(* Logix 5000 project; controller PLC_MCC1300_75F1 vendor 1 type 14 code 166 rev 32.11; software revision 32.04; part 64 of 83 *)
(* tags used below, declared in another part *)
   AUX_tConvoy_SL_NULL : UDT_Convoy_SL;
   CONST_rgdDestMask : DINT[32];   // Destination Mask
   CONST_tPlant : UDT_PLANT_CONSTANTS;
   GP_TrackingSearchPlate : GP_TrackingSearchPlate;
   M315Popup : MAC_Popup_ZC[2];
   M315Popup_HMW : MAC_Popup_ZC_HMW[2];
   M315Popup_ReentryCap : UDT_ConvoyCap_ZC;
   M315Popup_SL_DATA : UDT_Convoy_SL;
   M315Popup_tSearchPlateChangeFromCS4402 : GP_TrackingSearchPlate_STC;
   M315Popup_xDrivePosEnable : BOOL;
   M315Popup_xEndRise : BOOL;
   M315Popup_xEndRiseWaitingForCondition : BOOL;
   M350Popup : MAC_Popup_ZC;
   Sbr_INO_tConvoy_SL : UDT_Convoy_SL;
   TMP_d : DINT;
   TMP_dBaryc_ins_max : DINT;
   TMP_dBaryc_ins_min : DINT;
   TMP_dIndex : DINT;
   TMP_dIndexCap : DINT;
   TMP_dMaskAllowed : DINT;
   TMP_dStartSearch : DINT;
   TMP_dStopSearch : DINT;
   TMP_xAllCullet : BOOL;
   TMP_xAllLiteToCullet : BOOL;
   TMP_xAtLeastOneForSideLeg : BOOL;
   TMP_xDummy : BOOL;
   xAlwaysOFF : BOOL;
   Z300_BufferPlate : UDT_LINE_BUFFER_PLATE;
   Z300_Conveyor : UDT_StandConv[29];
   Z300_LineTracking : UDT_LINE_TRACKING;
   Z301 : MAC_Zone_ML;
(* MainProgram, continued *)

   // Rise request
   83: XIC(M315Popup[0].ST_xPlateInPositionToRise)[XIC(M315Popup[0].ST_xPlateToSinglePositioning) ,[XIC(M315Popup[0].ST_xPlateToBothPositioning) ,XIC(M315Popup[0].ST_xConvoyPositioning) ] [XIC(M315Popup[1].ST_xInitialConditionForRise) ,XIC(M315Popup[1].INPUT_xPopupHigh) ] ][XIC(M315Popup[0].ST_xInitialConditionForRise) ,XIC(M315Popup[0].INPUT_xPopupHigh) ,XIC(M315Popup[1].ST_xPlateToSinglePositioning) ][XIO(M315Popup[0].INPUT_xPopupHigh) XIO(M315Popup[1].ST_xPlateToSinglePositioning) XIO(Z300_Conveyor[26].OUTPUT_xPositioning.0) XIO(Z300_Conveyor[27].OUTPUT_xPositioning.0) XIO(Z300_Conveyor[28].OUTPUT_xPositioning.0) OTE(M315Popup[0].ST_xRequestRise) ,[XIC(M315Popup[0].ST_xPlateToBothPositioning) ,XIC(M315Popup[0].ST_xConvoyPositioning) ] XIO(M315Popup[1].INPUT_xPopupHigh) XIO(Z300_Conveyor[26].OUTPUT_xPositioning.0) XIO(Z300_Conveyor[27].OUTPUT_xPositioning.0) XIO(Z300_Conveyor[28].OUTPUT_xPositioning.0) OTE(M315Popup[1].ST_xRequestRise) ];
   // #####_Plate_ready_to_descend_#####
   84: JSR(sbrCheckConvoySLDestination,3,M315Popup_SL_DATA,M315Popup[0].AUX_dDestMaskOppOpSide,CONST_rgdDestMask[24],TMP_xAllCullet,TMP_xAtLeastOneForSideLeg);
   // #####_Descending_#####
   85: XIO(Z300_Conveyor[26].ST_xCleaningEnabled)LEQ(Z301.AUX_dBarPositionCleaning,970000)XIC(M315Popup[0].ST_xInitialConditionForDescend)XIO(M315Popup[0].ST_xPhasesInProgress)XIO(M315Popup[0].ST_xPlateUnderPopup)[XIO(M315Popup[0].ST_xPlatePresence) XIO(M315Popup[0].ST_xPlatePresentOnPopup) ,[XIC(M315Popup[0].ST_xPlatePresence) ,XIC(M315Popup[0].ST_xPlatePresentOnPopup) ] XIO(TMP_xAtLeastOneForSideLeg) ]XIO(Z300_LineTracking.rgtTrkConv[26].xGlassPresCom)XIO(Z300_LineTracking.rgtTrkConv[26].xGlassPresence)XIO(Z300_LineTracking.rgtTrkConv[27].xGlassPresCom)XIO(Z300_LineTracking.rgtTrkConv[27].xGlassPresence)XIO(M315Popup[0].INPUT_xPopupLow)XIO(M315Popup[0].tmOF_Wait.DN)XIO(Z300_Conveyor[26].OUTPUT_xPositioning.0)XIO(Z300_Conveyor[27].OUTPUT_xPositioning.0)XIO(Z300_Conveyor[28].OUTPUT_xPositioning.0)OTE(M315Popup[0].ST_xRequestDescend);
   // #####_Descending_#####
   86: XIO(Z300_Conveyor[26].ST_xCleaningEnabled)LEQ(Z301.AUX_dBarPositionCleaning,970000)XIC(M315Popup[1].ST_xInitialConditionForDescend)XIO(M315Popup[1].ST_xPhasesInProgress)XIO(M315Popup[1].ST_xPlateUnderPopup)[XIO(M315Popup[1].ST_xPlatePresence) XIO(M315Popup[1].ST_xPlatePresentOnPopup) ,[XIC(M315Popup[1].ST_xPlatePresence) ,XIC(M315Popup[1].ST_xPlatePresentOnPopup) ] ]XIO(Z300_LineTracking.rgtTrkConv[28].xGlassPresCom)XIO(Z300_LineTracking.rgtTrkConv[28].xGlassPresence)XIO(M315Popup[1].INPUT_xPopupLow)XIO(M315Popup[1].tmOF_Wait.DN)[XIO(Z300_Conveyor[26].OUTPUT_xPositioning.0) XIO(Z300_Conveyor[27].OUTPUT_xPositioning.0) ,XIO(xAlwaysOFF) ]XIO(Z300_Conveyor[28].OUTPUT_xPositioning.0)OTE(M315Popup[1].ST_xRequestDescend);
   87: [XIC(M315Popup[0].PH_xEndRise) ,XIC(M315Popup[1].PH_xEndRise) ]XIC(M315Popup_xEndRiseWaitingForCondition)OTE(M315Popup_xEndRise);
   88: [XIC(M315Popup[0].PH_xEndRise) ,XIC(M315Popup[1].PH_xEndRise) ,XIC(M315Popup_xEndRiseWaitingForCondition) ]OTE(M315Popup_xEndRiseWaitingForCondition);
   // #####_Move data to Popup_#####
   89: XIC(M315Popup[0].AUX_tSearchPlateData.xPlateHooked)XIC(M315Popup_xEndRise)[MOV(M315Popup[0].AUX_dIndexPositioning,TMP_dIndex) MOV(Z300_BufferPlate.rgtPlate[TMP_dIndex].tTracking.dPosition_cmm,M315Popup[0].AUX_dPosition_cmm) ,COP(AUX_tConvoy_SL_NULL,Sbr_INO_tConvoy_SL,1) ,JSR(sbrConvDataLineToSL,3,Z300_BufferPlate.rgtPlate[TMP_dIndex].tData,M315Popup_SL_DATA,0,Z300_BufferPlate.rgtPlate[TMP_dIndex].tData,M315Popup_SL_DATA) ,JSR(sbrConvDataLineToSL,3,Z300_BufferPlate.rgtPlate[TMP_dIndex].tData,M315Popup_SL_DATA,0,Z300_BufferPlate.rgtPlate[TMP_dIndex].tData,M315Popup_SL_DATA) ,MOV(0,M315Popup[0].AUX_dPosition_cmm) ,JSR(sbrTrackingDeleteConvoy,1,M315Popup[0].AUX_dIndexPositioning) ,OTU(M315Popup[0].AUX_tSearchPlateData.xPlateHooked) ,MOV(0,M315Popup[0].AUX_dIndexPositioning) ,MOV(0,M315Popup[0].AUX_dIndexPlatePositioned) ,OTL(M315Popup[0].ST_xPlatePresentOnPopup) ,OTU(M315Popup[0].ST_xPlateToBothPositioning) ,OTU(M315Popup[0].ST_xPlateToSinglePositioning) ,OTU(M315Popup[0].ST_xConvoyPositioning) ];
   90: XIC(M315Popup[0].ST_xPlatePresentOnPopup)OTE(M315Popup[0].ST_xPlateDataReadyToSend);
   91: XIC(M315Popup[1].ST_xPlatePresentOnPopup)OTE(M315Popup[1].ST_xPlateDataReadyToSend);
   92: ADD(Z300_LineTracking.rgtTrkConv[26].dStartPosition_cmm,310000,TMP_dBaryc_ins_min)SUB(Z300_LineTracking.rgtTrkConv[28].dEndPosition_cmm,310000,TMP_dBaryc_ins_max);
   // Convert from Convoy_ZLU to CapConvoy_ZC and Insert in tracking
   93: XIC(M315Popup[0].PH_xEndDescend)NEQ(M315Popup_SL_DATA.rgtCap[0].dID,0)[GRT(Z300_Conveyor[26].AUX_rgdTarget_cmm[0],0) ADD(Z300_LineTracking.rgtTrkConv[26].dStartPosition_cmm,Z300_Conveyor[26].AUX_rgdTarget_cmm[0],TMP_d) ,LEQ(Z300_Conveyor[26].AUX_rgdTarget_cmm[0],0) MOV(Z300_LineTracking.rgtTrkConv[28].dStartPosition_cmm,TMP_d) ]JSR(sbrResetLinkConvoy,0)JSR(sbrConvDataSLToLine,6,M315Popup_ReentryCap,M315Popup_SL_DATA,0,TMP_d,TMP_dBaryc_ins_min,TMP_dBaryc_ins_max,M315Popup_ReentryCap,M315Popup_SL_DATA)JSR(sbrPutLinkConvoy,0)JSR(sbrTrackingIndexTailConvoy,1,TMP_dIndex,M315Popup[0].AUX_dIndexPlateFree);
   // Delete plate data
   94: XIC(M315Popup[0].PH_xEndDescend)COP(AUX_tConvoy_SL_NULL,M315Popup_SL_DATA,1);
   95: XIO(M315Popup[0].ST_xPlateDataReadyToSend)XIC(M315Popup[0].INPUT_xPopupHigh)[XIC(M315Popup[0].ST_xPlatePresence) ,XIC(M315Popup[0].ST_xPlatePresentOnPopup) ]NEQ(M315Popup_SL_DATA.rgtCap[0].rgtLite[0].tDestination.rgxMain,CONST_rgdDestMask[24])ONS(M315Popup[0].OS_xPlateRemovedBySideLeg)[OTU(M315Popup[0].ST_xPlatePresence) ,COP(AUX_tConvoy_SL_NULL,M315Popup_SL_DATA,1) ,OTU(M315Popup[0].ST_xPlatePresentOnPopup) ];
   // #####_SATURATION_#####
   96: GRT(M315Popup_HMW[0].dSaturationSelection,0)XIC(Z301.ST_xCycleON)[[[XIC(Z300_LineTracking.rgtTrkConv[26].xGlassPresence) ,XIC(Z300_LineTracking.rgtTrkConv[27].xGlassPresence) ,XIC(Z300_LineTracking.rgtTrkConv[28].xGlassPresence) ,XIC(Z300_LineTracking.rgtTrkConv[26].xGlassPresCom) ,XIC(Z300_LineTracking.rgtTrkConv[27].xGlassPresCom) ,XIC(Z300_LineTracking.rgtTrkConv[28].xGlassPresCom) ] [XIO(Z300_Conveyor[26].ST_xRotationFeedback) ,XIO(Z300_Conveyor[27].ST_xRotationFeedback) ,XIO(Z300_Conveyor[28].ST_xRotationFeedback) ] ,XIO(xAlwaysOFF) [XIC(M315Popup[0].ST_xPlatePresence) XIC(M315Popup[0].INPUT_xPopupHigh) ,[XIO(M315Popup[0].ST_xInitialConditionForRise) ,XIO(M315Popup[1].ST_xInitialConditionForRise) ] ] ] ,LES(M315Popup_HMW[0].dSaturationSelection,1) ][[XIC(Z300_LineTracking.rgtTrkConv[25].xGlassPresence) ,XIC(Z300_LineTracking.rgtTrkConv[25].xGlassPresCom) ] XIO(Z300_Conveyor[25].ST_xRotationFeedback) ,LES(M315Popup_HMW[0].dSaturationSelection,2) ][[[XIC(Z300_LineTracking.rgtTrkConv[22].xGlassPresence) ,XIC(Z300_LineTracking.rgtTrkConv[23].xGlassPresence) ,XIC(Z300_LineTracking.rgtTrkConv[24].xGlassPresence) ,XIC(Z300_LineTracking.rgtTrkConv[22].xGlassPresCom) ,XIC(Z300_LineTracking.rgtTrkConv[23].xGlassPresCom) ,XIC(Z300_LineTracking.rgtTrkConv[24].xGlassPresCom) ] [XIO(Z300_Conveyor[22].ST_xRotationFeedback) ,XIO(Z300_Conveyor[23].ST_xRotationFeedback) ,XIO(Z300_Conveyor[24].ST_xRotationFeedback) ] ,XIC(M350Popup.INPUT_xPopupHigh) ] ,LES(M315Popup_HMW[0].dSaturationSelection,3) ][[XIC(Z300_LineTracking.rgtTrkConv[21].xGlassPresence) ,XIC(Z300_LineTracking.rgtTrkConv[21].xGlassPresCom) ] XIO(Z300_Conveyor[21].ST_xRotationFeedback) ,LES(M315Popup_HMW[0].dSaturationSelection,4) ][[XIC(Z300_LineTracking.rgtTrkConv[20].xGlassPresence) ,XIC(Z300_LineTracking.rgtTrkConv[20].xGlassPresCom) ] XIO(Z300_Conveyor[20].ST_xRotationFeedback) ,LES(M315Popup_HMW[0].dSaturationSelection,5) ]OTE(TMP_xDummy);
   97: XIC(TMP_xDummy)[[XIC(Z300_LineTracking.rgtTrkConv[19].xGlassPresence) ,XIC(Z300_LineTracking.rgtTrkConv[19].xGlassPresCom) ] XIO(Z300_Conveyor[19].ST_xRotationFeedback) ,LES(M315Popup_HMW[0].dSaturationSelection,6) ][[XIC(Z300_LineTracking.rgtTrkConv[18].xGlassPresence) ,XIC(Z300_LineTracking.rgtTrkConv[18].xGlassPresCom) ] XIO(Z300_Conveyor[18].ST_xRotationFeedback) ,LES(M315Popup_HMW[0].dSaturationSelection,7) ][[XIC(Z300_LineTracking.rgtTrkConv[17].xGlassPresence) ,XIC(Z300_LineTracking.rgtTrkConv[17].xGlassPresCom) ] XIO(Z300_Conveyor[17].ST_xRotationFeedback) ,LES(M315Popup_HMW[0].dSaturationSelection,8) ]OTE(TMP_xDummy);
   98: XIC(M315Popup[0].ST_xPlateComingToPopup)XIC(TMP_xDummy)[XIC(M315Popup[0].INPUT_xPopupHigh) ,XIO(xAlwaysOFF) [XIO(M315Popup[0].ST_xInitialConditionForRise) ,XIO(M315Popup[1].ST_xInitialConditionForRise) ] ][[XIO(M315Popup[0].ST_xInitialConditionForRise) ,XIO(M315Popup[1].ST_xInitialConditionForRise) ] [XIC(M315Popup[0].ST_xPlatePresence) ,XIO(xAlwaysOFF) [XIO(M315Popup[0].ST_xInitialConditionForRise) ,XIO(M315Popup[1].ST_xInitialConditionForRise) ] ] XIO(M315Popup[0].ST_xPlatePresentOnPopup) OTE(M315Popup[0].ST_xSaturationConditionPrevious) ,XIC(M315Popup[0].ST_xPlatePresentOnPopup) OTE(M315Popup[0].ST_xSaturationConditionPopup) ];
   99: XIC(M315Popup[0].ST_xPlateComingToPopup)XIC(TMP_xDummy)XIO(M315Popup_xEndRiseWaitingForCondition)XIC(M315Popup[0].INPUT_xPopupLow)XIO(M315Popup[0].ST_xPlatePresence)XIO(M315Popup[0].ST_xPlatePresentOnPopup)XIC(M315Popup[0].ST_xPlateStopToPopup)XIC(M315Popup[0].AUX_tSearchPlateData.xPlateHooked)NEQ(M315Popup[0].AUX_dIndexPositioning,0)OTE(M315Popup[0].ST_xSaturationConditionThis);
   100: GRT(M315Popup_HMW[0].dSaturationSelection,0)[XIC(M315Popup[0].ST_xSaturationConditionPrevious) XIO(M315Popup[0].ST_xSaturationConditionPopup) XIO(M315Popup[0].ST_xSaturationConditionThis) ,XIC(M315Popup[0].ST_xSaturationConditionThis) XIO(M315Popup[0].ST_xSaturationConditionPrevious) XIO(M315Popup[0].ST_xSaturationConditionPopup) ,XIC(M315Popup[0].ST_xSaturationConditionPopup) XIO(M315Popup[0].ST_xSaturationConditionPrevious) XIO(M315Popup[0].ST_xSaturationConditionThis) ]XIO(M315Popup[0].OS_xSaturationOnPrevious)XIO(M315Popup[0].OS_xSaturationOnThis)XIO(M315Popup[0].OS_xSaturationOnPopup)[XIO(Z300_Conveyor[23].OUTPUT_xPositioning.0) XIO(Z300_Conveyor[24].OUTPUT_xPositioning.0) ,XIO(Z300_Conveyor[22].ST_xRotationFeedback) XIO(M315Popup_xDrivePosEnable) ][XIO(M315Popup[0].ST_xRequestRise) XIO(M315Popup[1].ST_xRequestRise) ,XIO(M315Popup[0].ST_xInitialConditionForRise) ,XIO(M315Popup[1].ST_xInitialConditionForRise) ][TON(M315Popup[0].tmON_Saturation,?,?) ,XIC(M315Popup[0].tmON_Saturation.DN) [XIC(M315Popup[0].ST_xSaturationConditionPrevious) OTE(M315Popup[0].OS_xSaturationOnPrevious) ,XIC(M315Popup[0].ST_xSaturationConditionThis) OTE(M315Popup[0].OS_xSaturationOnThis) ,XIC(M315Popup[0].ST_xSaturationConditionPopup) OTE(M315Popup[0].OS_xSaturationOnPopup) ] ];
   // Allowed mask calculation for redestination
   101: CPT(TMP_dMaskAllowed,CONST_rgdDestMask[3]);
   102: XIC(M315Popup[0].OS_xSaturationOnPrevious)GRT(M315Popup[0].AUX_tSearchPlateData.dIndex,0)MOV(M315Popup[0].AUX_tSearchPlateData.dIndex,TMP_dIndexCap)[JSR(sbrRedestConvoyCapZC,5,M315Popup[0].AUX_tSearchPlateData.dIndex,M315Popup[0].AUX_dDestMaskOppOpSide,TMP_dMaskAllowed,0,CONST_rgdDestMask[24]) ,JSR(sbrTrackingIndexTailConvoy,1,M315Popup[0].AUX_tSearchPlateData.dIndex,M315Popup[0].AUX_dIndexPlateFree) ,[OTU(M315Popup[0].AUX_tSearchPlateData.xPlateHooked) ,MOV(0,M315Popup[0].AUX_dIndexPositioning) ] ];
   103: XIO(Z300_LineTracking.rgtTrkConv[25].xGlassPresence)XIO(Z300_LineTracking.rgtTrkConv[26].xGlassPresence)XIO(Z300_LineTracking.rgtTrkConv[27].xGlassPresence)XIO(Z300_LineTracking.rgtTrkConv[28].xGlassPresence)MOV(0,M315Popup[0].AUX_dIndexPlateFree);
   104: XIC(M315Popup[0].OS_xSaturationOnThis)XIC(M315Popup[0].AUX_tSearchPlateData.xPlateHooked)GRT(M315Popup[0].AUX_dIndexPlatePositioned,0)[JSR(sbrRedestConvoyCapZC,5,M315Popup[0].AUX_dIndexPlatePositioned,M315Popup[0].AUX_dDestMaskOppOpSide,TMP_dMaskAllowed,0,CONST_rgdDestMask[24]) ,OTU(M315Popup[0].AUX_tSearchPlateData.xPlateHooked) ,JSR(sbrTrackingIndexTailConvoy,1,M315Popup[0].AUX_dIndexPlatePositioned,M315Popup[0].AUX_dIndexPlateFree) ,MOV(0,M315Popup[0].AUX_dIndexPositioning) ,MOV(0,M315Popup[0].AUX_dIndexPlatePositioned) ];
   105: XIC(M315Popup[0].OS_xSaturationOnPopup)JSR(sbrRedestConvoySL,5,M315Popup_SL_DATA,M315Popup[0].AUX_dDestMaskOppOpSide,TMP_dMaskAllowed,0,CONST_rgdDestMask[24],M315Popup_SL_DATA);
   // Change destination of plate after popup if still has its destination
   106: ADD(150000,M315Popup[1].AUX_dEndPosition_cmm,TMP_dStartSearch)ADD(200000,M315Popup[1].AUX_dEndPosition_cmm,TMP_dStopSearch)GP_TrackingSearchPlate(GP_TrackingSearchPlate,TMP_dStartSearch,TMP_dStopSearch,0,Z300_LineTracking,M315Popup[0].tSearchPlateChangeDestAfterPopup,CONST_tPlant.dNumOfConveyors,CONST_tPlant.dNumCapsConveyor,Z300_BufferPlate);
   107: XIC(M315Popup[0].tSearchPlateChangeDestAfterPopup.xHeadPresence)ONS(M315Popup[0].OSR_xChangeDestAfterPopup)OTE(M315Popup[0].OS_xChangeDestAfterPopup);
   108: XIC(M315Popup[0].OS_xChangeDestAfterPopup)MOV(M315Popup[0].tSearchPlateChangeDestAfterPopup.rgdHeadPointer[0],M315Popup[0].AUX_dIndexPlateToChangeDestAfterPopup)CPT(TMP_dMaskAllowed,CONST_rgdDestMask[3])JSR(sbrRedestConvoyCapZC,5,M315Popup[0].tSearchPlateChangeDestAfterPopup.rgdHeadPointer,M315Popup[0].AUX_dDestMaskOppOpSide,TMP_dMaskAllowed,0,CONST_rgdDestMask[24]);
   // Change destination of plate if has its destination
   109: ADD(0,Z300_LineTracking.rgtTrkConv[25].dStartPosition_cmm,TMP_dStopSearch)ADD(0,Z300_LineTracking.rgtTrkConv[25].dEndPosition_cmm,TMP_dStartSearch)GP_TrackingSearchPlate(GP_TrackingSearchPlate,TMP_dStartSearch,TMP_dStopSearch,0,Z300_LineTracking,M315Popup_tSearchPlateChangeFromCS4402,CONST_tPlant.dNumOfConveyors,CONST_tPlant.dNumCapsConveyor,Z300_BufferPlate);
   // Verify destination
   110: GRT(M315Popup_tSearchPlateChangeFromCS4402.rgdHeadPointer[0],0)JSR(sbrCheckConvoyZCDestination,5,M315Popup_tSearchPlateChangeFromCS4402.rgdHeadPointer[0],M315Popup[0].AUX_dDestMaskOppOpSide,CONST_rgdDestMask[24],TMP_xAtLeastOneForSideLeg,TMP_xAllLiteToCullet,TMP_xAtLeastOneForSideLeg,TMP_xAllLiteToCullet);
   111: XIC(xAlwaysOFF)[XIC(M315Popup_tSearchPlateChangeFromCS4402.xHeadPresence) XIC(TMP_xAtLeastOneForSideLeg) MOV(CONST_rgdDestMask[3],TMP_dMaskAllowed) JSR(sbrRedestConvoyCapZC,5,M315Popup_tSearchPlateChangeFromCS4402.rgdHeadPointer,M315Popup[0].AUX_dDestMaskOppOpSide,TMP_dMaskAllowed,0,CONST_rgdDestMask[24]) ,XIC(M315Popup[0].AUX_tSearchPlateData.xPlateHooked) MOV(CONST_rgdDestMask[3],TMP_dMaskAllowed) JSR(sbrRedestConvoyCapZC,5,M315Popup[0].AUX_dIndexPositioning,M315Popup[0].AUX_dDestMaskOppOpSide,TMP_dMaskAllowed,0,CONST_rgdDestMask[24]) [OTU(M315Popup[0].AUX_tSearchPlateData.xPlateHooked) ,OTU(Z300_Conveyor[26].xReqPositioningHead) ,OTU(Z300_Conveyor[27].xReqPositioningHead) ,OTU(Z300_Conveyor[28].xReqPositioningHead) ,MOV(0,M315Popup[0].AUX_dIndexPositioning) ,MOV(0,M315Popup[0].AUX_dIndexPlatePositioned) ] ];
   // #####_CLEANING_#####
   112: XIC(Z300_Conveyor[26].ST_xCleaningEnabled)[OTU(M315Popup[0].PH_xRise) ,OTU(M315Popup[0].PH_xDescend) ,OTU(M315Popup[1].PH_xRise) ,OTU(M315Popup[1].PH_xDescend) ,MOV(0,M315Popup[0].AUX_dIndexPositioning) ,MOV(0,M315Popup[0].AUX_dIndexPlatePositioned) ,MOV(0,M315Popup[0].AUX_dIndexPlateFree) ,XIC(M315Popup[0].INPUT_xPopupLow) [COP(AUX_tConvoy_SL_NULL,M315Popup_SL_DATA,1) ,OTU(M315Popup[0].ST_xPlatePresence) ,OTU(M315Popup[0].ST_xPlatePresentOnPopup) ] ,XIC(M315Popup[1].INPUT_xPopupLow) [COP(AUX_tConvoy_SL_NULL,M315Popup_SL_DATA,1) ,OTU(M315Popup[1].ST_xPlatePresence) ,OTU(M315Popup[1].ST_xPlatePresentOnPopup) ] ];
   113: [XIC(M315Popup[0].INPUT_xPopupHigh) [COP(AUX_tConvoy_SL_NULL,M315Popup_SL_DATA,1) ,OTU(M315Popup[0].ST_xPlatePresence) ,OTU(M315Popup[0].ST_xPlatePresentOnPopup) ] ,XIC(M315Popup[1].INPUT_xPopupHigh) [COP(AUX_tConvoy_SL_NULL,M315Popup_SL_DATA,1) ,OTU(M315Popup[1].ST_xPlatePresence) ,OTU(M315Popup[1].ST_xPlatePresentOnPopup) ] ];
   114: XIO(M315Popup[0].AUX_tSearchPlateData.xPlateHooked)OTU(M315Popup[0].ST_xPlateToBothPositioning)OTU(M315Popup[0].ST_xPlateToSinglePositioning)OTU(M315Popup[1].ST_xPlateToSinglePositioning)OTU(M315Popup[0].ST_xConvoyPositioning);
END_ROUTINE
